   "DB_Displacement_Electromegnet" : Bool = PLC DB_Displacement.Electromagnet, 1 s
   "DB_HMI_Returning" : Bool = PLC DB_HMI.Returning, 100 ms

HMI tags "X_Axis"
   "DB_HMI_AxisStatus{0}_ActualPosition" : Real = PLC DB_HMI.AxisStatus[0].ActualPosition AT %DB1.DBW0, 500 ms
   "DB_HMI_AxisStatus{0}_ActualVelocity" : Real = PLC DB_HMI.AxisStatus[0].ActualVelocity AT %DB1.DBD0, 500 ms
   "DB_HMI_AxisStatus{0}_Error" : Bool = PLC DB_HMI.AxisStatus[0].Error AT %DB1.DBD0, 500 ms
   "DB_HMI_AxisStatus{0}_ErrorCode" : Word = PLC DB_HMI.AxisStatus[0].ErrorCode AT %DB1.DBX0.0, 500 ms
   "DB_HMI_AxisStatus{0}_Warning" : Bool = PLC DB_HMI.AxisStatus[0].Warning AT %DB1.DBX0.0, 500 ms
   "DB_HMI_AxisStatus{0}_WarningCode" : Word = PLC DB_HMI.AxisStatus[0].WarningCode AT %DB1.DBX0.0, 500 ms
   "DB_HMI_AxisStatus{0}_Referenced" : Bool = PLC DB_HMI.AxisStatus[0].Referenced AT %DB1.DBX0.0, 500 ms
   "DB_HMI_AxisStatus{0}_Enabled" : Bool = PLC DB_HMI.AxisStatus[0].Enabled AT %DB1.DBX0.0, 500 ms
   "DB_HMI_AxisStatus{0}_PositionReached" : Bool = PLC DB_HMI.AxisStatus[0].PositionReached AT %DB1.DBX0.0, 500 ms
   "DB_HMI_AxisControl{0}_JogActivate" : Bool = PLC DB_HMI.AxisControl[0].JogActivate AT %DB1.DBX0.0, 500 ms
   "DB_HMI_AxisControl{0}_JogCCW" : Bool = PLC DB_HMI.AxisControl[0].JogCCW AT %DB1.DBX0.0, 500 ms
   "DB_HMI_AxisControl{0}_JogCW" : Bool = PLC DB_HMI.AxisControl[0].JogCW AT %DB1.DBX0.0, 500 ms
   "DB_HMI_AxisControl{0}_ReqPosition" : Real = PLC DB_HMI.AxisControl[0].ReqPosition AT %DB1.DBX0.0, 500 ms
   "DB_HMI_AxisControl{0}_ReqVelocity" : Real = PLC DB_HMI.AxisControl[0].ReqVelocity AT %DB1.DBX0.0, 500 ms
   "DB_HMI_AxisControl{0}_SetReference" : Bool = PLC DB_HMI.AxisControl[0].SetReference AT %DB1.DBX0.0, 500 ms
   "DB_HMI_AxisControl{0}_Start" : Bool = PLC DB_HMI.AxisControl[0].Start AT %DB1.DBD0, 500 ms
   "DB_HMI_AxisControl{0}_Stop" : Bool = PLC DB_HMI.AxisControl[0].Stop AT %DB1.DBX0.0, 500 ms
   "DB_HMI_AxisStatus{0}_LimitCW" : Real = PLC DB_HMI.AxisStatus[0].LimitCW AT %DB1.DBW0, 500 ms
   "DB_HMI_AxisStatus{0}_LimitCCW" : Real = PLC DB_HMI.AxisStatus[0].LimitCCW AT %DB1.DBW0, 500 ms
   "DB_HMI_AxisStatus{0}_InvalidPosition" : Bool = PLC DB_HMI.AxisStatus[0].InvalidPosition AT %DB1.DBD0, 500 ms
   "DB_HMI_AxisStatus{0}_InvalidVelocity" : Bool = PLC DB_HMI.AxisStatus[0].InvalidVelocity AT %DB1.DBD0, 500 ms
   "DB_HMI_AxisStatus{0}_ParamCheckError" : Bool = PLC DB_HMI.AxisStatus[0].ParamCheckError AT %DB1.DBW0, 500 ms

HMI tags "Y_Axis"
   "DB_HMI_AxisStatus{1}_ActualPosition" : Real = PLC DB_HMI.AxisStatus[1].ActualPosition AT %DB1.DBW0, 500 ms
   "DB_HMI_AxisStatus{1}_ActualVelocity" : Real = PLC DB_HMI.AxisStatus[1].ActualVelocity AT %DB1.DBD0, 500 ms
   "DB_HMI_AxisStatus{1}_Error" : Bool = PLC DB_HMI.AxisStatus[1].Error AT %DB1.DBD0, 500 ms
   "DB_HMI_AxisStatus{1}_ErrorCode" : Word = PLC DB_HMI.AxisStatus[1].ErrorCode AT %DB1.DBX0.0, 500 ms
   "DB_HMI_AxisStatus{1}_Warning" : Bool = PLC DB_HMI.AxisStatus[1].Warning AT %DB1.DBX0.0, 500 ms
   "DB_HMI_AxisStatus{1}_WarningCode" : Word = PLC DB_HMI.AxisStatus[1].WarningCode AT %DB1.DBX0.0, 500 ms
   "DB_HMI_AxisStatus{1}_Referenced" : Bool = PLC DB_HMI.AxisStatus[1].Referenced AT %DB1.DBX0.0, 500 ms
   "DB_HMI_AxisStatus{1}_Enabled" : Bool = PLC DB_HMI.AxisStatus[1].Enabled AT %DB1.DBX0.0, 500 ms
   "DB_HMI_AxisStatus{1}_PositionReached" : Bool = PLC DB_HMI.AxisStatus[1].PositionReached AT %DB1.DBX0.0, 500 ms
   "DB_HMI_AxisControlAxisControl_1{1}_JogActivate" : Bool = PLC DB_HMI.AxisControl[1].JogActivate AT %DB1.DBX0.0, 500 ms
   "DB_HMI_AxisControlAxisControl_1{1}_JogCCW" : Bool = PLC DB_HMI.AxisControl[1].JogCCW AT %DB1.DBX0.0, 500 ms
   "DB_HMI_AxisControlAxisControl_1{1}_JogCW" : Bool = PLC DB_HMI.AxisControl[1].JogCW AT %DB1.DBX0.0, 500 ms
   "DB_HMI_AxisControlAxisControl_1{1}_ReqPosition" : Real = PLC DB_HMI.AxisControl[1].ReqPosition AT %DB1.DBX0.0, 500 ms
   "DB_HMI_AxisControlAxisControl_1{1}_ReqVelocity" : Real = PLC DB_HMI.AxisControl[1].ReqVelocity AT %DB1.DBX0.0, 500 ms
   "DB_HMI_AxisControlAxisControl_1{1}_SetReference" : Bool = PLC DB_HMI.AxisControl[1].SetReference AT %DB1.DBX0.0, 500 ms
   "DB_HMI_AxisControlAxisControl_1{1}_Start" : Bool = PLC DB_HMI.AxisControl[1].Start AT %DB1.DBD0, 500 ms
   "DB_HMI_AxisControlAxisControl_1{1}_Stop" : Bool = PLC DB_HMI.AxisControl[1].Stop AT %DB1.DBX0.0, 500 ms
   "DB_HMI_AxisStatus{1}_LimitCW" : Real = PLC DB_HMI.AxisStatus[1].LimitCW AT %DB1.DBW0, 500 ms
   "DB_HMI_AxisStatus{1}_LimitCCW" : Real = PLC DB_HMI.AxisStatus[1].LimitCCW AT %DB1.DBW0, 500 ms
   "DB_HMI_AxisStatus{1}_InvalidPosition" : Bool = PLC DB_HMI.AxisStatus[1].InvalidPosition AT %DB1.DBD0, 500 ms
   "DB_HMI_AxisStatus{1}_InvalidVelocity" : Bool = PLC DB_HMI.AxisStatus[1].InvalidVelocity AT %DB1.DBD0, 500 ms
   "DB_HMI_AxisStatus{1}_ParamCheckError" : Bool = PLC DB_HMI.AxisStatus[1].ParamCheckError AT %DB1.DBW0, 500 ms

HMI tags "Z_Axis"
   "DB_HMI_AxisStatus{2}_ActualPosition" : Real = PLC DB_HMI.AxisStatus[2].ActualPosition AT %DB1.DBW0, 500 ms
   "DB_HMI_AxisStatus{2}_ActualVelocity" : Real = PLC DB_HMI.AxisStatus[2].ActualVelocity AT %DB1.DBD0, 500 ms
   "DB_HMI_AxisStatus{2}_Error" : Bool = PLC DB_HMI.AxisStatus[2].Error AT %DB1.DBD0, 500 ms
   "DB_HMI_AxisStatus{2}_ErrorCode" : Word = PLC DB_HMI.AxisStatus[2].ErrorCode AT %DB1.DBX0.0, 500 ms
   "DB_HMI_AxisStatus{2}_Warning" : Bool = PLC DB_HMI.AxisStatus[2].Warning AT %DB1.DBX0.0, 500 ms
   "DB_HMI_AxisStatus{2}_WarningCode" : Word = PLC DB_HMI.AxisStatus[2].WarningCode AT %DB1.DBX0.0, 500 ms
   "DB_HMI_AxisStatus{2}_Referenced" : Bool = PLC DB_HMI.AxisStatus[2].Referenced AT %DB1.DBX0.0, 500 ms
   "DB_HMI_AxisStatus{2}_Enabled" : Bool = PLC DB_HMI.AxisStatus[2].Enabled AT %DB1.DBX0.0, 500 ms
   "DB_HMI_AxisStatus{2}_PositionReached" : Bool = PLC DB_HMI.AxisStatus[2].PositionReached AT %DB1.DBX0.0, 500 ms
   "DB_HMI_AxisControlAxisControl{2}_JogActivate" : Bool = PLC DB_HMI.AxisControl[2].JogActivate AT %DB1.DBX0.0, 500 ms
   "DB_HMI_AxisControlAxisControl{2}_JogCCW" : Bool = PLC DB_HMI.AxisControl[2].JogCCW AT %DB1.DBX0.0, 500 ms
   "DB_HMI_AxisControlAxisControl{2}_JogCW" : Bool = PLC DB_HMI.AxisControl[2].JogCW AT %DB1.DBX0.0, 500 ms
   "DB_HMI_AxisControlAxisControl{2}_ReqPosition" : Real = PLC DB_HMI.AxisControl[2].ReqPosition AT %DB1.DBX0.0, 500 ms
   "DB_HMI_AxisControlAxisControl{2}_ReqVelocity" : Real = PLC DB_HMI.AxisControl[2].ReqVelocity AT %DB1.DBX0.0, 500 ms
   "DB_HMI_AxisControlAxisControl{2}_SetReference" : Bool = PLC DB_HMI.AxisControl[2].SetReference AT %DB1.DBX0.0, 500 ms
   "DB_HMI_AxisControlAxisControl{2}_Start" : Bool = PLC DB_HMI.AxisControl[2].Start AT %DB1.DBD0, 500 ms
   "DB_HMI_AxisControlAxisControl{2}_Stop" : Bool = PLC DB_HMI.AxisControl[2].Stop AT %DB1.DBX0.0, 500 ms
   "DB_HMI_AxisStatus{2}_LimitCW" : Real = PLC DB_HMI.AxisStatus[2].LimitCW AT %DB1.DBW0, 500 ms
   "DB_HMI_AxisStatus{2}_LimitCCW" : Real = PLC DB_HMI.AxisStatus[2].LimitCCW AT %DB1.DBW0, 500 ms
   "DB_HMI_AxisStatus{2}_InvalidPosition" : Bool = PLC DB_HMI.AxisStatus[2].InvalidPosition AT %DB1.DBD0, 500 ms
   "DB_HMI_AxisStatus{2}_InvalidVelocity" : Bool = PLC DB_HMI.AxisStatus[2].InvalidVelocity AT %DB1.DBD0, 500 ms
   "DB_HMI_AxisStatus{2}_ParamCheckError" : Bool = PLC DB_HMI.AxisStatus[2].ParamCheckError AT %DB1.DBW0, 500 ms

HMI tags "Electromagnet"
   "Electromagnet" : Bool = PLC Electromagnet AT %Q8.0, 500 ms
   "Laser_Sensor" : Bool = PLC Laser_Sensor AT %I8.5, 100 ms

HMI tags "Sensors"
   "Inductive_Sensor_4" : Bool = PLC Inductive_Sensor_4 AT %I8.0, 500 ms
   "Inductive_Sensor_3" : Bool = PLC Inductive_Sensor_3 AT %I8.1, 500 ms
   "Inductive_Sensor_2" : Bool = PLC Inductive_Sensor_2 AT %I8.2, 500 ms
   "Inductive_Sensor_1" : Bool = PLC Inductive_Sensor_1 AT %I8.3, 500 ms

screen "Main" 800x480, template "Template_1"
   on GenerateScreen: SetTag("ScreenNumber", 1)
   TextField "Text field_1" at 16,187 size 764x82; Text 'Stanowisko Pozycjoner'
   TextField "Text field_7" at 149,0 size 552x50; Text 'Main Screen'
   Circle "Circle_1" at 31,367 size 31x31
      Appearance <- "DB_HMI_Interrupt"
   Button "Button_3" at 588,360 size 192x50; TextOff 'Searching'
      on Click: ActivateScreen("Searching", 0)

Template "Template_1" 800x480
   Group "Group" at 0,0 size 800x50; Picture "Graphic_13"
   Button "Button_2" at 0,428 size 100x52; TextOff 'Main Screen'
      on Click: ActivateScreen("Main", 0)
      Appearance <- "ScreenNumber"
   Button "Button_4" at 100,428 size 100x52; TextOff 'X Axis'
      on Click: ActivateScreen("X_Axis", 0)
      Appearance <- "ScreenNumber"
   Button "Button_3" at 300,428 size 100x52; TextOff 'Z Axis'
      on Click: ActivateScreen("Z_Axis", 0)
      Appearance <- "ScreenNumber"
   Button "Button_5" at 400,428 size 100x52; TextOff 'Electro- magnet'
      on Click: ActivateScreen("Electromagnet", 0)
      Appearance <- "ScreenNumber"
   Button "Button_6" at 500,428 size 100x52; TextOff 'Sensors'
      Appearance <- "ScreenNumber"
      on Click: ActivateScreen("Sensors", 0)
   Button "Button_7" at 600,428 size 100x52; TextOff 'Enable'
      on Press: SetBit("DB_HMI_Enable")
      Appearance <- "DB_HMI_Enable"
      on Release: ResetBit("DB_HMI_Enable")
   Button "Button_8" at 700,428 size 100x52; TextOff 'Reset'
      on Release: ResetBit("DB_HMI_Reset")
      on Press: SetBit("DB_HMI_Reset")
      Appearance <- "DB_HMI_Reset"
   Button "Button_9" at 200,428 size 100x52; TextOff 'Y Axis'
      on Click: ActivateScreen("Y_Axis", 0)
      Appearance <- "ScreenNumber"
   Rectangle "Rectangle_9" at 700,0 size 100x50
      Appearance <- "EStop_Fdb"
   TextField "Text field_2" at 721,14 size 59x23; Text 'E-Stop'
   GraphicView "Template_Graphic view_1" at 2,2 size 146x46; Picture "Graphic_13"

screen "X_Axis" 800x480, template "Template_1"
   on ClearScreen: ResetBit("DB_HMI_AxisControl{0}_JogActivate")
   on GenerateScreen: SetTag("ScreenNumber", 2)
   TextField "Text field_3" at 23,204 size 42x29; Text 'Jog'
   TextField "Text field_4" at 22,68 size 109x29; Text 'Reference'
   TextField "Text field_6" at 269,68 size 152x29; Text 'Go to position'
   Group "Group_2" at 265,67 size 341x219
   Group "Group_1" at 19,203 size 240x130
   Group "Group" at 19,67 size 240x130
   Button "Button_3" at 88,219 size 100x50; TextOff 'Activate'
      on Click: InvertBit("DB_HMI_AxisControl{0}_JogActivate")
      Appearance <- "DB_HMI_AxisControl{0}_JogActivate"
   Button "Button_4" at 26,276 size 100x50; TextOff 'Jog REV'
      on Release: ResetBit("DB_HMI_AxisControl{0}_JogCW")
      on Press: SetBit("DB_HMI_AxisControl{0}_JogCW")
      Appearance <- "DB_HMI_AxisControl{0}_JogCW"
   Button "Button_5" at 150,276 size 100x50; TextOff 'Jog FW'
      on Release: ResetBit("DB_HMI_AxisControl{0}_JogCCW")
      on Press: SetBit("DB_HMI_AxisControl{0}_JogCCW")
      Appearance <- "DB_HMI_AxisControl{0}_JogCCW"
   IOField "I/O field_1" at 387,127 size 108x50; FormatPattern 9999.9; Unit mm
      ProcessValue <- "DB_HMI_AxisControl{0}_ReqPosition"
   IOField "I/O field_2" at 387,215 size 108x50; FormatPattern 999; Unit mm/s
      ProcessValue <- "DB_HMI_AxisControl{0}_ReqVelocity"
   TextField "Text field_1" at 268,140 size 119x23; Text 'Req. Position:'
   TextField "Text field_2" at 268,228 size 118x23; Text 'Req. Velocity:'
   Button "Button_6" at 499,127 size 100x50; TextOff 'Start'
      on Release: ResetBit("DB_HMI_AxisControl{0}_Start")
      on Press: SetBit("DB_HMI_AxisControl{0}_Start")
   Circle "Circle_1" at 25,103 size 24x24
      Appearance <- "DB_HMI_AxisStatus{0}_Referenced"
   TextField "Text field_5" at 51,104 size 146x23; Text 'Drive Referenced'
   Button "Button_1" at 89,140 size 100x50; TextOff 'Set Reference'
      on Release: ResetBit("DB_HMI_AxisControl{0}_SetReference")
      on Press: SetBit("DB_HMI_AxisControl{0}_SetReference")
   Button "Button_2" at 499,215 size 100x50; TextOff 'Stop'
      on Release: ResetBit("DB_HMI_AxisControl{0}_Stop")
      on Press: SetBit("DB_HMI_AxisControl{0}_Stop")
   TextField "Text field_8" at 616,68 size 106x29; Text 'Drive info'
   Circle "Circle_2" at 620,103 size 24x24
      Appearance <- "DB_HMI_AxisStatus{0}_Enabled"
   TextField "Text field_9" at 646,104 size 118x23; Text 'Drive Enabled'
   TextField "Text field_10" at 646,133 size 146x23; Text 'Position Reached'
   Circle "Circle_3" at 620,132 size 24x24
      Appearance <- "DB_HMI_AxisStatus{0}_PositionReached"
   Circle "Circle_4" at 620,277 size 24x24
      Appearance <- "DB_HMI_AxisStatus{0}_Warning"
   TextField "Text field_11" at 646,278 size 73x23; Text 'Warning'
   TextField "Text field_12" at 620,307 size 105x23; Text 'Warn. Code:'
   IOField "I/O field_4" at 702,162 size 90x23; FormatPattern 9999.9; Unit mm
      ProcessValue <- "DB_HMI_AxisStatus{0}_ActualPosition"
   IOField "I/O field_5" at 699,191 size 100x23; FormatPattern s999; Unit mm/s
      ProcessValue <- "DB_HMI_AxisStatus{0}_ActualVelocity"
   TextField "Text field_13" at 620,162 size 77x23; Text 'Position:'
   TextField "Text field_14" at 620,191 size 76x23; Text 'Velocity:'
   TextField "Text field_15" at 620,220 size 84x23; Text 'CW Limit:'
   TextField "Text field_16" at 620,249 size 95x23; Text 'CCW Limit:'
   IOField "I/O field_6" at 715,220 size 80x23; FormatPattern 999; Unit mm
      ProcessValue <- "DB_HMI_AxisStatus{0}_LimitCW"
   IOField "I/O field_7" at 715,249 size 80x23; FormatPattern 9999; Unit mm
      ProcessValue <- "DB_HMI_AxisStatus{0}_LimitCCW"
   IOField "I/O field_3" at 729,307 size 60x23; FormatPattern 99999
      ProcessValue <- "DB_HMI_AxisStatus{0}_WarningCode"
   Circle "Circle_5" at 620,336 size 24x24
      Appearance <- "DB_HMI_AxisStatus{0}_Error"
   TextField "Text field_17" at 646,337 size 46x23; Text 'Error'
   TextField "Text field_18" at 620,366 size 98x23; Text 'Error Code:'
   IOField "I/O field_8" at 728,366 size 60x23; FormatPattern 99999
      ProcessValue <- "DB_HMI_AxisStatus{0}_ErrorCode"
   Circle "Circle_6" at 273,103 size 24x24
      Appearance <- "DB_HMI_AxisStatus{0}_InvalidPosition"
   TextField "Text field_19" at 299,104 size 224x23; Text 'Invalid Requested Position'
   Circle "Circle_7" at 273,191 size 24x24
      Appearance <- "DB_HMI_AxisStatus{0}_InvalidVelocity"
   TextField "Text field_20" at 299,192 size 223x23; Text 'Invalid Requested Velocity'
   Circle "Circle_8" at 620,395 size 24x24
      Appearance <- "DB_HMI_AxisStatus{0}_ParamCheckError"
   TextField "Text field_21" at 646,396 size 138x23; Text 'Error Parameter'
   TextField "Text field_7" at 149,0 size 552x50; Text 'X Axis'

screen "Y_Axis" 800x480, template "Template_1"
   on GenerateScreen: SetTag("ScreenNumber", 3)
   on ClearScreen: ResetBit("DB_HMI_AxisControlAxisControl_1{1}_JogActivate")
   TextField "Text field_3" at 23,204 size 42x29; Text 'Jog'
   TextField "Text field_4" at 22,68 size 109x29; Text 'Reference'
   TextField "Text field_6" at 269,68 size 152x29; Text 'Go to position'
   Group "Group_2" at 265,67 size 341x219
   Group "Group_1" at 19,203 size 240x130
   Group "Group" at 19,67 size 240x130
   Button "Button_3" at 88,219 size 100x50; TextOff 'Activate'
      on Click: InvertBit("DB_HMI_AxisControlAxisControl_1{1}_JogActivate")
      Appearance <- "DB_HMI_AxisControlAxisControl_1{1}_JogActivate"
   Button "Button_4" at 26,276 size 100x50; TextOff 'Jog REV'
      on Release: ResetBit("DB_HMI_AxisControlAxisControl_1{1}_JogCW")
      on Press: SetBit("DB_HMI_AxisControlAxisControl_1{1}_JogCW")
      Appearance <- "DB_HMI_AxisControlAxisControl_1{1}_JogCW"
   Button "Button_5" at 150,276 size 100x50; TextOff 'Jog FW'
      on Release: ResetBit("DB_HMI_AxisControlAxisControl_1{1}_JogCCW")
      on Press: SetBit("DB_HMI_AxisControlAxisControl_1{1}_JogCCW")
      Appearance <- "DB_HMI_AxisControlAxisControl_1{1}_JogCCW"
   Circle "Circle_1" at 25,103 size 24x24
      Appearance <- "DB_HMI_AxisStatus{1}_Referenced"
   TextField "Text field_5" at 51,104 size 146x23; Text 'Drive Referenced'
   Button "Button_1" at 89,140 size 100x50; TextOff 'Set Reference'
      on Release: ResetBit("DB_HMI_AxisControlAxisControl_1{1}_SetReference")
      on Press: SetBit("DB_HMI_AxisControlAxisControl_1{1}_SetReference")
   TextField "Text field_8" at 616,68 size 106x29; Text 'Drive info'
   Circle "Circle_2" at 620,103 size 24x24
      Appearance <- "DB_HMI_AxisStatus{1}_Enabled"
   TextField "Text field_9" at 646,104 size 118x23; Text 'Drive Enabled'
   TextField "Text field_10" at 646,133 size 146x23; Text 'Position Reached'
   Circle "Circle_3" at 620,132 size 24x24
      Appearance <- "DB_HMI_AxisStatus{1}_PositionReached"
   Circle "Circle_4" at 620,277 size 24x24
      Appearance <- "DB_HMI_AxisStatus{1}_Warning"
   TextField "Text field_11" at 646,278 size 73x23; Text 'Warning'
   TextField "Text field_12" at 620,307 size 105x23; Text 'Warn. Code:'
   TextField "Text field_13" at 620,162 size 77x23; Text 'Position:'
   TextField "Text field_14" at 620,191 size 76x23; Text 'Velocity:'
   TextField "Text field_15" at 620,220 size 84x23; Text 'CW Limit:'
   TextField "Text field_16" at 620,249 size 95x23; Text 'CCW Limit:'
   IOField "I/O field_3" at 729,307 size 60x23; FormatPattern 99999
      ProcessValue <- "DB_HMI_AxisStatus{1}_WarningCode"
   Circle "Circle_5" at 620,336 size 24x24
      Appearance <- "DB_HMI_AxisStatus{1}_Error"
   TextField "Text field_17" at 646,337 size 46x23; Text 'Error'
   TextField "Text field_18" at 620,366 size 98x23; Text 'Error Code:'
   IOField "I/O field_8" at 728,366 size 60x23; FormatPattern 99999
      ProcessValue <- "DB_HMI_AxisStatus{1}_ErrorCode"
   IOField "I/O field_5" at 699,191 size 100x23; FormatPattern s999; Unit mm/s
      ProcessValue <- "DB_HMI_AxisStatus{1}_ActualVelocity"
   IOField "I/O field_6" at 715,220 size 80x23; FormatPattern 999; Unit mm
      ProcessValue <- "DB_HMI_AxisStatus{1}_LimitCW"
   IOField "I/O field_7" at 715,249 size 80x23; FormatPattern 9999; Unit mm
      ProcessValue <- "DB_HMI_AxisStatus{1}_LimitCCW"
   TextField "Text field_1" at 268,140 size 119x23; Text 'Req. Position:'
   TextField "Text field_2" at 268,228 size 118x23; Text 'Req. Velocity:'
   Button "Button_6" at 499,127 size 100x50; TextOff 'Start'
      on Release: ResetBit("DB_HMI_AxisControlAxisControl_1{1}_Start")
      on Press: SetBit("DB_HMI_AxisControlAxisControl_1{1}_Start")
   Button "Button_2" at 499,215 size 100x50; TextOff 'Stop'
      on Release: ResetBit("DB_HMI_AxisControlAxisControl_1{1}_Stop")
      on Press: SetBit("DB_HMI_AxisControlAxisControl_1{1}_Stop")
   IOField "I/O field_1" at 387,127 size 108x50; FormatPattern 9999.9; Unit mm
      ProcessValue <- "DB_HMI_AxisControlAxisControl_1{1}_ReqPosition"
   IOField "I/O field_2" at 387,215 size 108x50; FormatPattern 999; Unit mm/s
      ProcessValue <- "DB_HMI_AxisControlAxisControl_1{1}_ReqVelocity"
   Circle "Circle_6" at 273,103 size 24x24
      Appearance <- "DB_HMI_AxisStatus{1}_InvalidPosition"
   TextField "Text field_19" at 299,104 size 224x23; Text 'Invalid Requested Position'
   Circle "Circle_7" at 273,191 size 24x24
      Appearance <- "DB_HMI_AxisStatus{1}_InvalidVelocity"
   TextField "Text field_20" at 299,192 size 223x23; Text 'Invalid Requested Velocity'
   IOField "I/O field_4" at 702,162 size 90x23; FormatPattern 9999.9; Unit mm
      ProcessValue <- "DB_HMI_AxisStatus{1}_ActualPosition"
   Circle "Circle_8" at 620,395 size 24x24
      Appearance <- "DB_HMI_AxisStatus{1}_ParamCheckError"
   TextField "Text field_21" at 646,396 size 138x23; Text 'Error Parameter'
   TextField "Text field_7" at 149,0 size 552x50; Text 'Y Axis'

screen "Z_Axis" 800x480, template "Template_1"
   on GenerateScreen: SetTag("ScreenNumber", 4)
   on ClearScreen: ResetBit("DB_HMI_AxisControlAxisControl{2}_JogActivate")
   TextField "Text field_3" at 23,204 size 42x29; Text 'Jog'
   TextField "Text field_4" at 22,68 size 109x29; Text 'Reference'
   TextField "Text field_6" at 269,68 size 152x29; Text 'Go to position'
   Group "Group_2" at 265,67 size 341x219
   Group "Group_1" at 19,203 size 240x130
   Group "Group" at 19,67 size 240x130
   Button "Button_3" at 88,219 size 100x50; TextOff 'Activate'
      on Click: InvertBit("DB_HMI_AxisControlAxisControl{2}_JogActivate")
      Appearance <- "DB_HMI_AxisControlAxisControl{2}_JogActivate"
   Button "Button_4" at 26,276 size 100x50; TextOff 'Jog REV'
      on Release: ResetBit("DB_HMI_AxisControlAxisControl{2}_JogCW")
      on Press: SetBit("DB_HMI_AxisControlAxisControl{2}_JogCW")
      Appearance <- "DB_HMI_AxisControlAxisControl{2}_JogCW"
   Button "Button_5" at 150,276 size 100x50; TextOff 'Jog FW'
      on Release: ResetBit("DB_HMI_AxisControlAxisControl{2}_JogCCW")
      on Press: SetBit("DB_HMI_AxisControlAxisControl{2}_JogCCW")
      Appearance <- "DB_HMI_AxisControlAxisControl{2}_JogCCW"
   Circle "Circle_1" at 25,103 size 24x24
      Appearance <- "DB_HMI_AxisStatus{2}_Referenced"
   TextField "Text field_5" at 51,104 size 146x23; Text 'Drive Referenced'
   Button "Button_1" at 89,140 size 100x50; TextOff 'Set Reference'
      on Release: ResetBit("DB_HMI_AxisControlAxisControl{2}_SetReference")
      on Press: SetBit("DB_HMI_AxisControlAxisControl{2}_SetReference")
   TextField "Text field_8" at 616,68 size 106x29; Text 'Drive info'
   Circle "Circle_2" at 620,103 size 24x24
      Appearance <- "DB_HMI_AxisStatus{2}_Enabled"
   TextField "Text field_9" at 646,104 size 118x23; Text 'Drive Enabled'
   TextField "Text field_10" at 646,133 size 146x23; Text 'Position Reached'
   Circle "Circle_3" at 620,132 size 24x24
      Appearance <- "DB_HMI_AxisStatus{2}_PositionReached"
   Circle "Circle_4" at 620,277 size 24x24
      Appearance <- "DB_HMI_AxisStatus{2}_Warning"
   TextField "Text field_11" at 646,278 size 73x23; Text 'Warning'
   TextField "Text field_12" at 620,307 size 105x23; Text 'Warn. Code:'
   TextField "Text field_13" at 620,162 size 77x23; Text 'Position:'
   TextField "Text field_14" at 620,191 size 76x23; Text 'Velocity:'
   TextField "Text field_15" at 620,220 size 84x23; Text 'CW Limit:'
   TextField "Text field_16" at 620,249 size 95x23; Text 'CCW Limit:'
   IOField "I/O field_3" at 729,307 size 60x23; FormatPattern 99999
      ProcessValue <- "DB_HMI_AxisStatus{2}_WarningCode"
   Circle "Circle_5" at 620,336 size 24x24
      Appearance <- "DB_HMI_AxisStatus{2}_Error"
   TextField "Text field_17" at 646,337 size 46x23; Text 'Error'
   TextField "Text field_18" at 620,366 size 98x23; Text 'Error Code:'
   IOField "I/O field_8" at 728,366 size 60x23; FormatPattern 99999
      ProcessValue <- "DB_HMI_AxisStatus{2}_ErrorCode"
   IOField "I/O field_5" at 699,191 size 100x23; FormatPattern s999; Unit mm/s
      ProcessValue <- "DB_HMI_AxisStatus{2}_ActualVelocity"
   TextField "Text field_1" at 268,140 size 119x23; Text 'Req. Position:'
   TextField "Text field_2" at 268,228 size 118x23; Text 'Req. Velocity:'
   Button "Button_6" at 499,127 size 100x50; TextOff 'Start'
      on Release: ResetBit("DB_HMI_AxisControlAxisControl{2}_Start")
      on Press: SetBit("DB_HMI_AxisControlAxisControl{2}_Start")
   Button "Button_2" at 499,215 size 100x50; TextOff 'Stop'
      on Release: ResetBit("DB_HMI_AxisControlAxisControl{2}_Stop")
      on Press: SetBit("DB_HMI_AxisControlAxisControl{2}_Stop")
   IOField "I/O field_1" at 387,127 size 108x50; FormatPattern 9999.9; Unit mm
      ProcessValue <- "DB_HMI_AxisControlAxisControl{2}_ReqPosition"
   IOField "I/O field_2" at 387,215 size 108x50; FormatPattern 999; Unit mm/s
      ProcessValue <- "DB_HMI_AxisControlAxisControl{2}_ReqVelocity"
   IOField "I/O field_6" at 715,220 size 80x23; FormatPattern 999; Unit mm
      ProcessValue <- "DB_HMI_AxisStatus{2}_LimitCW"
   IOField "I/O field_7" at 715,249 size 80x23; FormatPattern 9999; Unit mm
      ProcessValue <- "DB_HMI_AxisStatus{2}_LimitCCW"
   Circle "Circle_6" at 273,103 size 24x24
      Appearance <- "DB_HMI_AxisStatus{2}_InvalidPosition"
   TextField "Text field_19" at 299,104 size 224x23; Text 'Invalid Requested Position'
   Circle "Circle_7" at 273,191 size 24x24
      Appearance <- "DB_HMI_AxisStatus{2}_InvalidVelocity"
   TextField "Text field_20" at 299,192 size 223x23; Text 'Invalid Requested Velocity'
   IOField "I/O field_4" at 702,162 size 90x23; FormatPattern 9999.9; Unit mm
      ProcessValue <- "DB_HMI_AxisStatus{2}_ActualPosition"
   Circle "Circle_8" at 620,395 size 24x24
      Appearance <- "DB_HMI_AxisStatus{2}_ParamCheckError"
   TextField "Text field_21" at 646,396 size 138x23; Text 'Error Parameter'
   TextField "Text field_7" at 149,0 size 552x50; Text 'Z Axis'

screen "Electromagnet" 800x480, template "Template_1"
   on GenerateScreen: SetTag("ScreenNumber", 5)
   TextField "Text field_3" at 22,204 size 189x29; Text 'Electromagnet L1'
   Group "Group_1" at 19,203 size 204x112
   Group "Group" at 19,67 size 204x104
   Button "Button_3" at 71,245 size 100x50; TextOff 'Activate'
      on Click: InvertBit("DB_HMI_Electromagnet")
      Appearance <- "Electromagnet"
   Circle "Circle_1" at 25,115 size 24x24
      Appearance <- "Laser Sensor"
   TextField "Text field_5" at 51,116 size 119x23; Text 'Part Detected'
   TextField "Text field_7" at 149,0 size 552x50; Text 'Electromagnet'
   TextField "Text field_4" at 22,68 size 172x29; Text 'Laser Sensor A1'

screen "Sensors" 800x480, template "Template_1"
   on GenerateScreen: SetTag("ScreenNumber", 6)
   TextField "Text field_4" at 21,68 size 160x29; Text 'Part Sensor B1'
   Group "Group" at 19,67 size 166x104
   Circle "Circle_1" at 25,115 size 24x24
      Appearance <- "Inductive_Sensor_1"
   TextField "Text field_5" at 51,116 size 119x23; Text 'Part Detected'
   Group "Group_1" at 217,67 size 166x104
   Group "Group_2" at 415,67 size 166x104
   Group "Group_3" at 613,67 size 166x104
   Circle "Circle_2" at 223,115 size 24x24
      Appearance <- "Inductive_Sensor_2"
   TextField "Text field_6" at 249,116 size 119x23; Text 'Part Detected'
   Circle "Circle_3" at 421,115 size 24x24
      Appearance <- "Inductive_Sensor_3"
   TextField "Text field_7" at 447,116 size 119x23; Text 'Part Detected'
   Circle "Circle_4" at 619,115 size 24x24
      Appearance <- "Inductive_Sensor_4"
   TextField "Text field_8" at 645,116 size 119x23; Text 'Part Detected'
   TextField "Text field_9" at 149,0 size 552x50; Text 'Sensors'
   TextField "Text field_1" at 219,68 size 160x29; Text 'Part Sensor B2'
   TextField "Text field_2" at 417,68 size 160x29; Text 'Part Sensor B3'
   TextField "Text field_3" at 615,68 size 160x29; Text 'Part Sensor B4'

screen "Searching" 800x480
   Button "Button_1" at 45,12 size 121x42; TextOff 'Searching'
      on Press: InvertBit("DB_HMI_Searching"); ResetBit("DB_HMI_StartPosition")
      Appearance <- "DB_HMI_Searching"
   Button "Button_2" at 188,12 size 133x41; TextOff 'Start position'
      on Press: InvertBit("DB_HMI_StartPosition"); ResetBit("DB_HMI_Searching")
      Appearance <- "DB_HMI_StartPosition"
   Button "Button_3" at 661,15 size 97x42; TextOff 'Main'
      on Click: ActivateScreen("Main", 0)
   TextField "Text field_31" at 315,431 size 124x23; Text 'Electromagnet'
   Circle "Circle_4" at 450,428 size 34x34
      Appearance <- "DB_Displacement_Electromegnet"
   TextField "Text field_32" at 550,325 size 136x23; Text 'Active Interrupt'
   Circle "Circle_5" at 697,317 size 34x34
      Appearance <- "Drivers_Interrupt_DB_Interrupt_Active"
   Group "Group" at 550,367 size 181x98
   Group "Group_1" at 11,70 size 248x225
   Group "Group_2" at 270,70 size 248x225
   Group "Group_3" at 529,70 size 248x226
   Group "Group_4" at 308,312 size 201x104
   Group "Group_5" at 7,313 size 280x75
   Group "Group_6" at 20,394 size 220x80
   Button "Button_6" at 427,320 size 74x32; TextOff 'Reset'
      on Press: SetBit("DB_HMI_ResetSpace")
      on Release: ResetBit("DB_HMI_ResetSpace")
   Button "Button_7" at 321,366 size 38x37; TextOff 'Text'
      on Press: InvertBit("DB_HMI_PlaceOcc_S1"); InvertBit("DB_Displacement_PlaceOcup_Sens1")
      Appearance <- "DB_Displacement_PlaceOcup_Sens1"
   Button "Button_8" at 369,367 size 36x37; TextOff 'Text'
      on Press: InvertBit("DB_HMI_PlaceOcc_S2"); InvertBit("DB_Displacement_PlaceOcup_Sens2")
      Appearance <- "DB_Displacement_PlaceOcup_Sens2"
   Button "Button_9" at 413,367 size 34x37; TextOff 'Text'
      on Press: InvertBit("DB_HMI_PlaceOcc_S3"); InvertBit("DB_Displacement_PlaceOcup_Sens3")
      Appearance <- "DB_Displacement_PlaceOcup_Sens3"
   Button "Button_10" at 457,367 size 37x37; TextOff 'Text'
      on Press: InvertBit("DB_HMI_PlaceOcc_S4"); InvertBit("DB_Displacement_PlaceOcup_Sens4")
      Appearance <- "DB_Displacement_PlaceOcup_Sens4"
   TextField "Text field_40" at 19,358 size 254x23; Text 'Return to the starting position'
      Visibility <- "DB_HMI_Returning"
   TextField "Text field_41" at 82,358 size 131x23; Text 'Invalid position'
      Visibility <- "DB_HMI_ErrorState"
   Button "Button_11" at 148,401 size 69x30; TextOff 'Reset'
      Visibility <- "DB_HMI_ErrorState"
   Button "Button_12" at 148,436 size 69x31; TextOff 'Enable'
      Visibility <- "DB_HMI_ErrorState"
   TextField "Text field_1" at 23,78 size 56x23; Text 'Axis X'
   TextField "Text field_2" at 46,112 size 71x23; Text 'Position'
   TextField "Text field_3" at 45,141 size 70x23; Text 'Velocity'
   TextField "Text field_4" at 45,173 size 78x23; Text 'Limit CW'
   TextField "Text field_5" at 46,205 size 89x23; Text 'Limit CCW'
   TextField "Text field_6" at 46,248 size 46x23; Text 'Error'
   IOField "I/O field_1" at 147,109 size 96x32; FormatPattern s999999999.999
      ProcessValue <- "Drivers_DB_UDT_Axis_Status{0}_ActualPosition"
   IOField "I/O field_2" at 147,138 size 96x32; FormatPattern s999999999.999
      ProcessValue <- "Drivers_DB_UDT_Axis_Status{0}_ActualVelocity"
   IOField "I/O field_3" at 147,165 size 96x32; FormatPattern s999999999.999
      ProcessValue <- "Drivers_DB_UDT_Axis_Status{0}_LimitCW"
   IOField "I/O field_4" at 147,193 size 96x32; FormatPattern s999999999.999
      ProcessValue <- "Drivers_DB_UDT_Axis_Status{0}_LimitCCW"
   Circle "Circle_1" at 181,248 size 34x34
      Appearance <- "FB_Axis_X_DB_o_Status_Error"
   IOField "I/O field_5" at 405,116 size 96x32; FormatPattern s999999999.999
      ProcessValue <- "FB_Axis_Y_DB_o_Status_ActualPosition"
   IOField "I/O field_6" at 405,144 size 96x32; FormatPattern s999999999.999
      ProcessValue <- "FB_Axis_Y_DB_o_Status_ActualVelocity"
   IOField "I/O field_7" at 405,172 size 96x32; FormatPattern s999999999.999
      ProcessValue <- "FB_Axis_Y_DB_o_Status_LimitCW"
   IOField "I/O field_8" at 405,199 size 96x32; FormatPattern s999999999.999
      ProcessValue <- "FB_Axis_Y_DB_o_Status_LimitCCW"
   TextField "Text field_7" at 279,75 size 56x23; Text 'Axis Y'
   TextField "Text field_8" at 302,109 size 71x23; Text 'Position'
   TextField "Text field_9" at 301,138 size 70x23; Text 'Velocity'
   TextField "Text field_10" at 301,170 size 78x23; Text 'Limit CW'
   TextField "Text field_11" at 302,202 size 89x23; Text 'Limit CCW'
   TextField "Text field_12" at 302,245 size 46x23; Text 'Error'
   Circle "Circle_2" at 442,248 size 34x34
      Appearance <- "FB_Axis_Y_DB_o_Status_Error"
   IOField "I/O field_9" at 662,112 size 96x32; FormatPattern s999999999.999
      ProcessValue <- "FB_Axis_Z_DB_o_Status_ActualPosition"
   IOField "I/O field_10" at 662,140 size 96x32; FormatPattern s999999999.999
      ProcessValue <- "FB_Axis_Z_DB_o_Status_ActualVelocity"
   IOField "I/O field_11" at 662,167 size 96x32; FormatPattern s999999999.999
      ProcessValue <- "FB_Axis_Z_DB_o_Status_LimitCW"
   IOField "I/O field_12" at 662,196 size 96x32; FormatPattern s999999999.999
      ProcessValue <- "FB_Axis_Z_DB_o_Status_LimitCCW"
   TextField "Text field_13" at 535,72 size 55x23; Text 'Axis Z'
   TextField "Text field_14" at 558,106 size 71x23; Text 'Position'
   TextField "Text field_15" at 557,135 size 70x23; Text 'Velocity'
   TextField "Text field_16" at 557,167 size 78x23; Text 'Limit CW'
   TextField "Text field_17" at 558,199 size 89x23; Text 'Limit CCW'
   TextField "Text field_18" at 558,242 size 46x23; Text 'Error'
   Circle "Circle_3" at 698,248 size 34x34
      Appearance <- "FB_Axis_Z_DB_o_Status_Error"
   TextField "Text field_19" at 24,316 size 114x23; Text 'Actual Status'
   TextField "Text field_20" at 66,358 size 155x23; Text 'Searching for item'
      Visibility <- "Interrupts_DB_GeneralCounter"
   TextField "Text field_21" at 78,357 size 132x23; Text 'Item was found'
      Visibility <- "DB_HMI_ItemwasFound"
   TextField "Text field_22" at 41,355 size 200x23; Text 'Center point calculation'
      Visibility <- "DB_HMI_MidPosCounting"
   TextField "Text field_23" at 65,358 size 153x23; Text 'Grabbing the item'
      Visibility <- "DB_HMI_GrabbingTheItem"
   TextField "Text field_24" at 26,357 size 234x23; Text 'The item has been set aside'
      Visibility <- "DB_Displacement_Electromegnet"
   TextField "Text field_35" at 68,358 size 157x23; Text 'No space available'
      Visibility <- "DB_HMI_AvailablePlace"
   TextField "Text field_37" at 29,357 size 231x23; Text 'Moving to the start position'
      Visibility <- "DB_HMI_MovingToStartPosition"
   TextField "Text field_38" at 46,358 size 192x23; Text 'Start Position Reached'
      Visibility <- "DB_HMI_StartPositionReached"
   TextField "Text field_25" at 327,332 size 68x23; Text 'Sensors'
   TextField "Text field_26" at 320,317 size 81x23; Text 'Inductive'
   Rectangle "Rectangle_6" at 323,366 size 34x37
      Appearance <- "DB_Displacement_PlaceOcup_Sens1"
   TextField "Text field_27" at 333,374 size 15x23; Text '1'
   Rectangle "Rectangle_7" at 369,366 size 34x37
      Appearance <- "DB_Displacement_PlaceOcup_Sens2"
   TextField "Text field_28" at 379,374 size 15x23; Text '2'
   Rectangle "Rectangle_8" at 413,366 size 34x37
      Appearance <- "DB_Displacement_PlaceOcup_Sens3"
   TextField "Text field_29" at 423,374 size 15x23; Text '3'
   Rectangle "Rectangle_9" at 459,366 size 34x37
      Appearance <- "DB_Displacement_PlaceOcup_Sens4"
   TextField "Text field_30" at 469,374 size 15x23; Text '4'
   TextField "Text field_33" at 554,402 size 56x23; Text 'X AVG'
   TextField "Text field_34" at 553,428 size 56x23; Text 'Y AVG'
   IOField "I/O field_13" at 629,399 size 96x32; FormatPattern s999999999.999
      ProcessValue <- "Drivers_DB_X_AVG"
   IOField "I/O field_14" at 629,426 size 96x32; FormatPattern s999999999.999
      ProcessValue <- "Drivers_DB_Y_AVG"
   TextField "Text field_39" at 580,368 size 108x23; Text 'Center Point'
   Circle "Circle_6" at 93,418 size 34x34
      Appearance <- "DB_HMI_ErrorState"
   TextField "Text field_36" at 42,423 size 46x23; Text 'Error'
   Button "Button_4" at 147,401 size 69x31; TextOff 'Reset'
      Appearance <- "DB_HMI_ResetError"
      on Release: ResetBit("DB_HMI_ResetError")
      on Press: SetBit("DB_HMI_ResetError")
      Visibility <- "DB_HMI_ErrorState"
   Button "Button_5" at 147,436 size 69x31; TextOff 'Enable'
      on Press: SetBit("DB_HMI_Start/Enable")
      on Release: ResetBit("DB_HMI_Start/Enable")
      Appearance <- "DB_HMI_Start/Enable"
      Visibility <- "DB_HMI_ErrorState"
*)